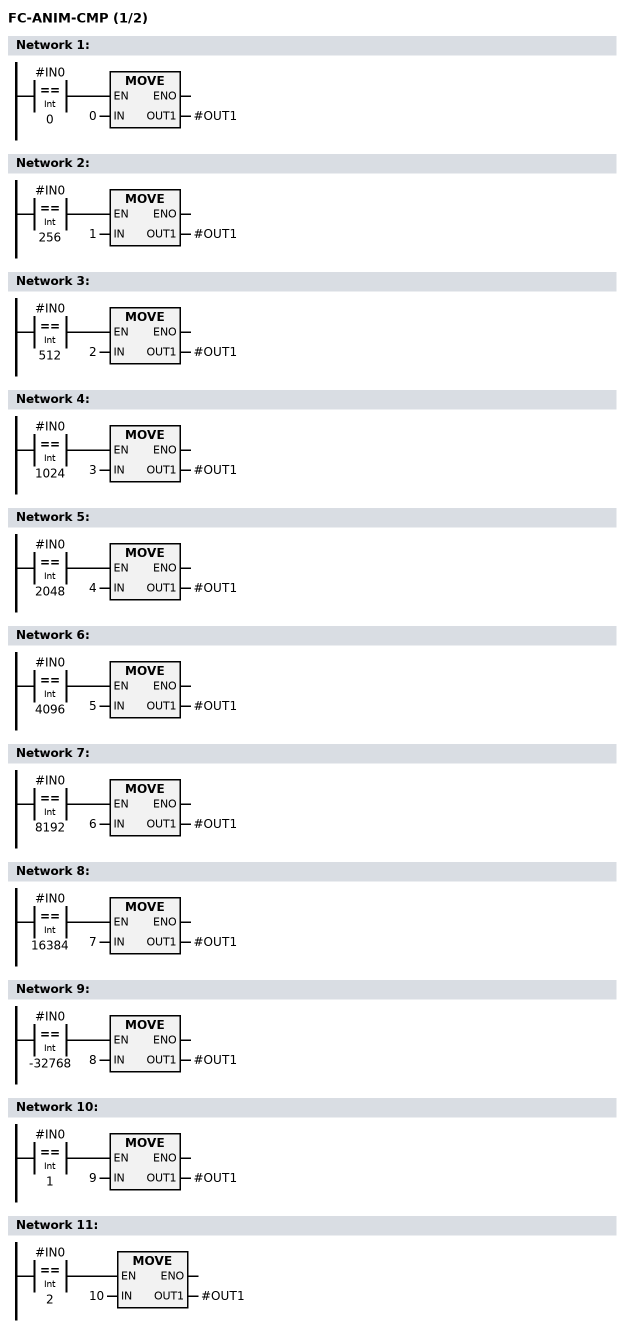
   RUNG wire#powerrail
      { S7_Templates := "SrcType := Int" } EQ_Contact(in1 := #IN0, in2 := 0)
      { S7_GenerateENO := "TRUE" } Move(in := 0, out1 => #OUT1)
   END_RUNG
   // the same network as SCL:
   IF #IN0 = 0 THEN #OUT1 := 0; END_IF;
END_REGION

REGION Network 2
   RUNG wire#powerrail
      { S7_Templates := "SrcType := Int" } EQ_Contact(in1 := #IN0, in2 := 256)
      { S7_GenerateENO := "TRUE" } Move(in := 1, out1 => #OUT1)
   END_RUNG
   // the same network as SCL:
   IF #IN0 = 256 THEN #OUT1 := 1; END_IF;
END_REGION

REGION Network 3
   RUNG wire#powerrail
      { S7_Templates := "SrcType := Int" } EQ_Contact(in1 := #IN0, in2 := 512)
      { S7_GenerateENO := "TRUE" } Move(in := 2, out1 => #OUT1)
   END_RUNG
   // the same network as SCL:
   IF #IN0 = 512 THEN #OUT1 := 2; END_IF;
END_REGION

REGION Network 4
   RUNG wire#powerrail
      { S7_Templates := "SrcType := Int" } EQ_Contact(in1 := #IN0, in2 := 1024)
      { S7_GenerateENO := "TRUE" } Move(in := 3, out1 => #OUT1)
   END_RUNG
   // the same network as SCL:
   IF #IN0 = 1024 THEN #OUT1 := 3; END_IF;
END_REGION

REGION Network 5
   RUNG wire#powerrail
      { S7_Templates := "SrcType := Int" } EQ_Contact(in1 := #IN0, in2 := 2048)
      { S7_GenerateENO := "TRUE" } Move(in := 4, out1 => #OUT1)
   END_RUNG
   // the same network as SCL:
   IF #IN0 = 2048 THEN #OUT1 := 4; END_IF;
END_REGION

REGION Network 6
   RUNG wire#powerrail
      { S7_Templates := "SrcType := Int" } EQ_Contact(in1 := #IN0, in2 := 4096)
      { S7_GenerateENO := "TRUE" } Move(in := 5, out1 => #OUT1)
   END_RUNG
   // the same network as SCL:
   IF #IN0 = 4096 THEN #OUT1 := 5; END_IF;
END_REGION

REGION Network 7
   RUNG wire#powerrail
      { S7_Templates := "SrcType := Int" } EQ_Contact(in1 := #IN0, in2 := 8192)
      { S7_GenerateENO := "TRUE" } Move(in := 6, out1 => #OUT1)
   END_RUNG
   // the same network as SCL:
   IF #IN0 = 8192 THEN #OUT1 := 6; END_IF;
END_REGION

REGION Network 8
   RUNG wire#powerrail
      { S7_Templates := "SrcType := Int" } EQ_Contact(in1 := #IN0, in2 := 16384)
      { S7_GenerateENO := "TRUE" } Move(in := 7, out1 => #OUT1)
   END_RUNG
   // the same network as SCL:
   IF #IN0 = 16384 THEN #OUT1 := 7; END_IF;
END_REGION

REGION Network 9
   RUNG wire#powerrail
      { S7_Templates := "SrcType := Int" } EQ_Contact(in1 := #IN0, in2 := -32768)
      { S7_GenerateENO := "TRUE" } Move(in := 8, out1 => #OUT1)
   END_RUNG
   // the same network as SCL:
   IF #IN0 = (-32768) THEN #OUT1 := 8; END_IF;
END_REGION

REGION Network 10
   RUNG wire#powerrail
      { S7_Templates := "SrcType := Int" } EQ_Contact(in1 := #IN0, in2 := 1)
      { S7_GenerateENO := "TRUE" } Move(in := 9, out1 => #OUT1)
   END_RUNG
   // the same network as SCL:
   IF #IN0 = 1 THEN #OUT1 := 9; END_IF;
END_REGION

REGION Network 11
   RUNG wire#powerrail
      { S7_Templates := "SrcType := Int" } EQ_Contact(in1 := #IN0, in2 := 2)
      { S7_GenerateENO := "TRUE" } Move(in := 10, out1 => #OUT1)
   END_RUNG
   // the same network as SCL:
   IF #IN0 = 2 THEN #OUT1 := 10; END_IF;
END_REGION

REGION Network 12
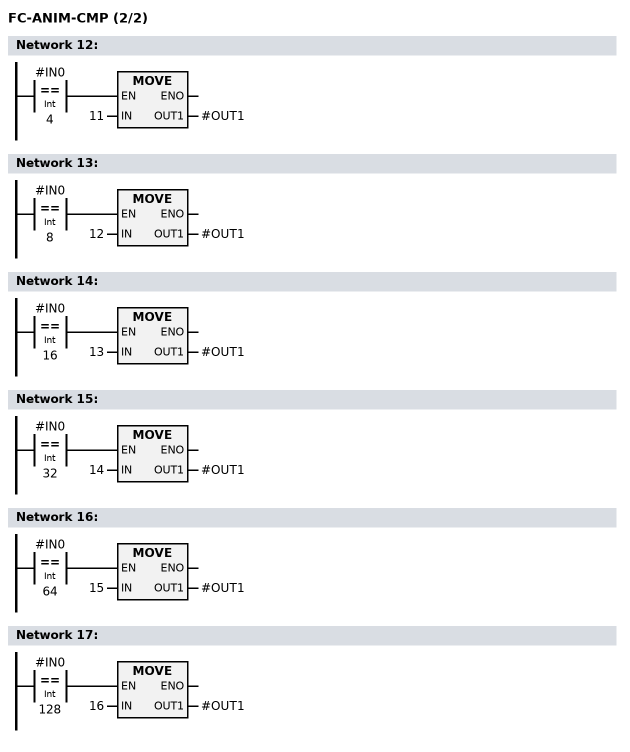
   RUNG wire#powerrail
      { S7_Templates := "SrcType := Int" } EQ_Contact(in1 := #IN0, in2 := 4)
      { S7_GenerateENO := "TRUE" } Move(in := 11, out1 => #OUT1)
   END_RUNG
   // the same network as SCL:
   IF #IN0 = 4 THEN #OUT1 := 11; END_IF;
END_REGION

REGION Network 13
   RUNG wire#powerrail
      { S7_Templates := "SrcType := Int" } EQ_Contact(in1 := #IN0, in2 := 8)
      { S7_GenerateENO := "TRUE" } Move(in := 12, out1 => #OUT1)
   END_RUNG
   // the same network as SCL:
   IF #IN0 = 8 THEN #OUT1 := 12; END_IF;
END_REGION

REGION Network 14
   RUNG wire#powerrail
      { S7_Templates := "SrcType := Int" } EQ_Contact(in1 := #IN0, in2 := 16)
      { S7_GenerateENO := "TRUE" } Move(in := 13, out1 => #OUT1)
   END_RUNG
   // the same network as SCL:
   IF #IN0 = 16 THEN #OUT1 := 13; END_IF;
END_REGION

REGION Network 15
   RUNG wire#powerrail
      { S7_Templates := "SrcType := Int" } EQ_Contact(in1 := #IN0, in2 := 32)
      { S7_GenerateENO := "TRUE" } Move(in := 14, out1 => #OUT1)
   END_RUNG
   // the same network as SCL:
   IF #IN0 = 32 THEN #OUT1 := 14; END_IF;
END_REGION

REGION Network 16
   RUNG wire#powerrail
      { S7_Templates := "SrcType := Int" } EQ_Contact(in1 := #IN0, in2 := 64)
      { S7_GenerateENO := "TRUE" } Move(in := 15, out1 => #OUT1)
   END_RUNG
   // the same network as SCL:
   IF #IN0 = 64 THEN #OUT1 := 15; END_IF;
END_REGION

REGION Network 17
   RUNG wire#powerrail
      { S7_Templates := "SrcType := Int" } EQ_Contact(in1 := #IN0, in2 := 128)
      { S7_GenerateENO := "TRUE" } Move(in := 16, out1 => #OUT1)
   END_RUNG
   // the same network as SCL:
   IF #IN0 = 128 THEN #OUT1 := 16; END_IF;
END_REGION
END_FUNCTION

// folder: Panel/Iluminación

FUNCTION "IluminaciónMTA" : Void   // FC23, LAD
{ S7_Optimized_Access := 'FALSE' }
VERSION : 0.1
// LUC - 05/08/2020
   VAR_TEMP   // added for the SCL form of the ladder/FBD networks
      _s5time1 : S5Time;
   END_VAR
BEGIN

REGION Network 1: Seteo de temporizador desde panel
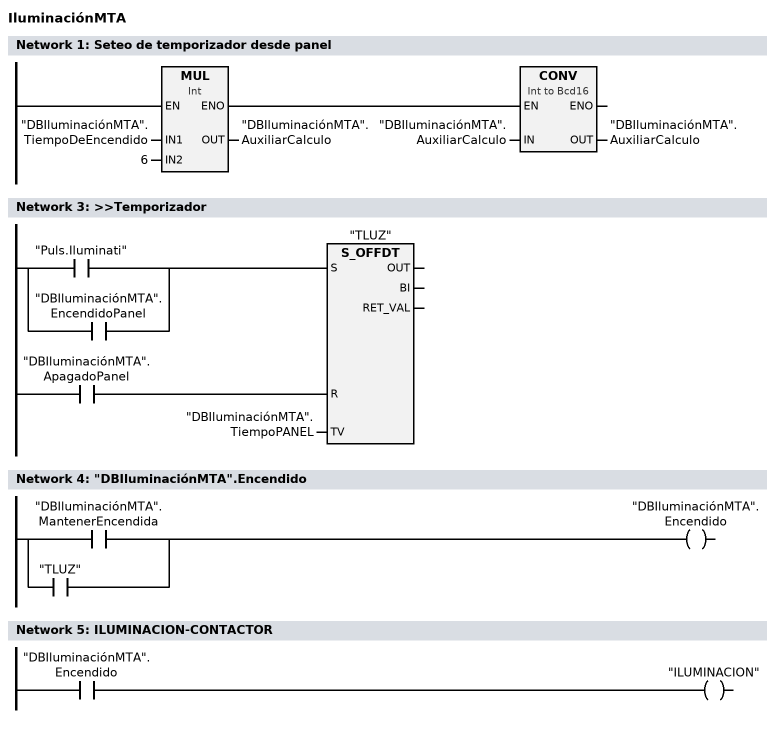
   RUNG wire#powerrail
      { S7_Templates := "SrcType := Int"; S7_GenerateENO := "TRUE" } Mul(in1 := "DBIluminaciónMTA".TiempoDeEncendido, in2 := 6, out => "DBIluminaciónMTA".AuxiliarCalculo)
      { S7_Templates := "[SrcType := Int, DestType := Bcd16]"; S7_GenerateENO := "TRUE" } Convert(in := "DBIluminaciónMTA".AuxiliarCalculo, out => "DBIluminaciónMTA".AuxiliarCalculo)
   END_RUNG
   // the same network as SCL:
   // ENO of a box is taken as its EN; it also drops when the box reports an error
   "DBIluminaciónMTA".AuxiliarCalculo := "DBIluminaciónMTA".TiempoDeEncendido * 6;
   "DBIluminaciónMTA".AuxiliarCalculo := INT_TO_BCD16("DBIluminaciónMTA".AuxiliarCalculo);
END_REGION

REGION Network 2 (STL): Seteo de temporizador desde panel
         L     12288;
         L     "DBIluminaciónMTA".AuxiliarCalculo;
         OW;
         T     "DBIluminaciónMTA".TiempoPANEL;
         NOP   0;
END_REGION

REGION Network 3: >>Temporizador
   RUNG wire#powerrail
      Contact( "Puls.Iluminati" )
      wire#w1
      S_OFFDT(T_NO := "TLUZ", R := wire#w2, TV := "DBIluminaciónMTA".TiempoPANEL, BI =>, RET_VAL =>)
   END_RUNG
   RUNG wire#powerrail
      Contact( "DBIluminaciónMTA".EncendidoPanel )
   END_RUNG wire#w1
   RUNG wire#powerrail
      Contact( "DBIluminaciónMTA".ApagadoPanel )
   END_RUNG wire#w2
   // the same network as SCL:
   #_s5time1 := S_OFFDT(T_NO := "TLUZ",
                        S := "Puls.Iluminati" OR "DBIluminaciónMTA".EncendidoPanel,
                        R := "DBIluminaciónMTA".ApagadoPanel,
                        TV := "DBIluminaciónMTA".TiempoPANEL);
END_REGION

REGION Network 4: "DBIluminaciónMTA".Encendido
   RUNG wire#powerrail
      Contact( "DBIluminaciónMTA".MantenerEncendida )
      wire#w1
      Coil( "DBIluminaciónMTA".Encendido )
   END_RUNG
   RUNG wire#powerrail
      Contact( "TLUZ" )
   END_RUNG wire#w1
   // the same network as SCL:
   "DBIluminaciónMTA".Encendido := "DBIluminaciónMTA".MantenerEncendida OR "TLUZ";
END_REGION

REGION Network 5: ILUMINACION-CONTACTOR
   RUNG wire#powerrail
      Contact( "DBIluminaciónMTA".Encendido )
      Coil( "ILUMINACION" )
   END_RUNG
   // the same network as SCL:
   "ILUMINACION" := "DBIluminaciónMTA".Encendido;
END_REGION
END_FUNCTION

// folder: Secadores/Alta

FUNCTION "EnclavSecAltaMTA" : Void   // FC12, LAD
{ S7_Optimized_Access := 'FALSE' }
VERSION : 0.1
BEGIN

REGION Network 1: Arranque automático MS050
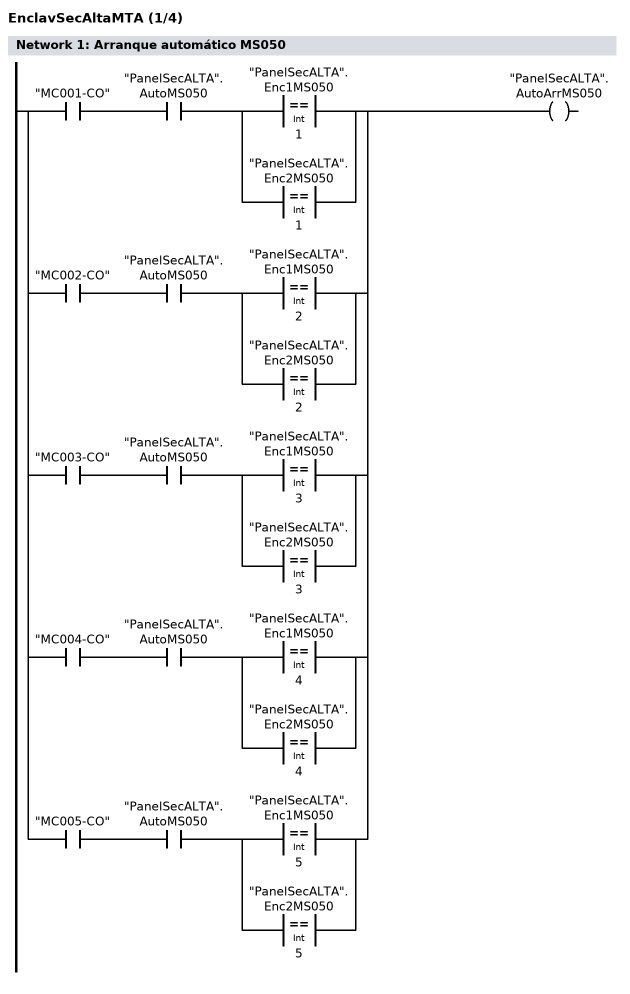
   RUNG wire#powerrail
      Contact( "MC001-CO" )
      Contact( "PanelSecALTA".AutoMS050 )
      wire#w1
      { S7_Templates := "SrcType := Int" } EQ_Contact(in1 := "PanelSecALTA".Enc1MS050, in2 := 1)
      wire#w2
      Coil( "PanelSecALTA".AutoArrMS050 )
   END_RUNG
   RUNG wire#w1
      { S7_Templates := "SrcType := Int" } EQ_Contact(in1 := "PanelSecALTA".Enc2MS050, in2 := 1)
   END_RUNG wire#w2
   RUNG wire#powerrail
      Contact( "MC002-CO" )
      Contact( "PanelSecALTA".AutoMS050 )
      wire#w3
      { S7_Templates := "SrcType := Int" } EQ_Contact(in1 := "PanelSecALTA".Enc1MS050, in2 := 2)
   END_RUNG wire#w2
   RUNG wire#w3
      { S7_Templates := "SrcType := Int" } EQ_Contact(in1 := "PanelSecALTA".Enc2MS050, in2 := 2)
   END_RUNG wire#w2
   RUNG wire#powerrail
      Contact( "MC003-CO" )
      Contact( "PanelSecALTA".AutoMS050 )
      wire#w4
      { S7_Templates := "SrcType := Int" } EQ_Contact(in1 := "PanelSecALTA".Enc1MS050, in2 := 3)
   END_RUNG wire#w2
   RUNG wire#w4
      { S7_Templates := "SrcType := Int" } EQ_Contact(in1 := "PanelSecALTA".Enc2MS050, in2 := 3)
   END_RUNG wire#w2
   RUNG wire#powerrail
      Contact( "MC004-CO" )
      Contact( "PanelSecALTA".AutoMS050 )
      wire#w5
      { S7_Templates := "SrcType := Int" } EQ_Contact(in1 := "PanelSecALTA".Enc1MS050, in2 := 4)
   END_RUNG wire#w2
   RUNG wire#w5
      { S7_Templates := "SrcType := Int" } EQ_Contact(in1 := "PanelSecALTA".Enc2MS050, in2 := 4)
   END_RUNG wire#w2
   RUNG wire#powerrail
      Contact( "MC005-CO" )
      Contact( "PanelSecALTA".AutoMS050 )
      wire#w6
      { S7_Templates := "SrcType := Int" } EQ_Contact(in1 := "PanelSecALTA".Enc1MS050, in2 := 5)
   END_RUNG wire#w2
   RUNG wire#w6
      { S7_Templates := "SrcType := Int" } EQ_Contact(in1 := "PanelSecALTA".Enc2MS050, in2 := 5)
   END_RUNG wire#w2
   // the same network as SCL:
   "PanelSecALTA".AutoArrMS050 := ("MC001-CO" AND "PanelSecALTA".AutoMS050 AND (("PanelSecALTA".Enc1MS050 = 1) OR ("PanelSecALTA".Enc2MS050 = 1))) OR ("MC002-CO" AND "PanelSecALTA".AutoMS050 AND (("PanelSecALTA".Enc1MS050 = 2) OR ("PanelSecALTA".Enc2MS050 = 2))) OR ("MC003-CO" AND "PanelSecALTA".AutoMS050 AND (("PanelSecALTA".Enc1MS050 = 3) OR ("PanelSecALTA".Enc2MS050 = 3))) OR ("MC004-CO" AND "PanelSecALTA".AutoMS050 AND (("PanelSecALTA".Enc1MS050 = 4) OR ("PanelSecALTA".Enc2MS050 = 4))) OR ("MC005-CO" AND "PanelSecALTA".AutoMS050 AND (("PanelSecALTA".Enc1MS050 = 5) OR ("PanelSecALTA".Enc2MS050 = 5)));
END_REGION

REGION Network 2: Arranque automático MS051
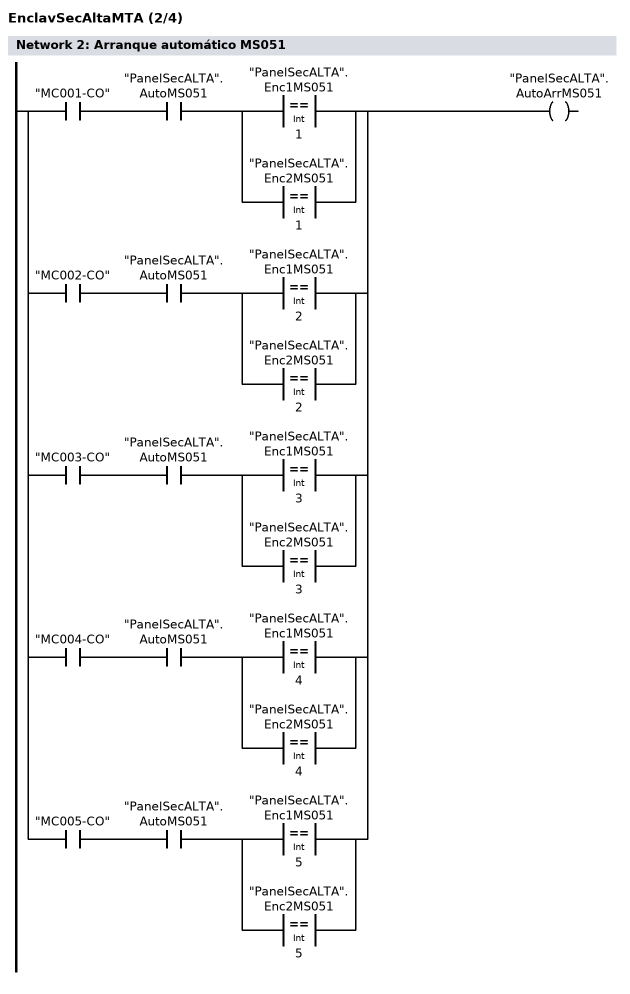
   RUNG wire#powerrail
      Contact( "MC001-CO" )
      Contact( "PanelSecALTA".AutoMS051 )
      wire#w1
      { S7_Templates := "SrcType := Int" } EQ_Contact(in1 := "PanelSecALTA".Enc1MS051, in2 := 1)
      wire#w2
      Coil( "PanelSecALTA".AutoArrMS051 )
   END_RUNG
   RUNG wire#w1
      { S7_Templates := "SrcType := Int" } EQ_Contact(in1 := "PanelSecALTA".Enc2MS051, in2 := 1)
   END_RUNG wire#w2
   RUNG wire#powerrail
      Contact( "MC002-CO" )
      Contact( "PanelSecALTA".AutoMS051 )
      wire#w3
      { S7_Templates := "SrcType := Int" } EQ_Contact(in1 := "PanelSecALTA".Enc1MS051, in2 := 2)
   END_RUNG wire#w2
   RUNG wire#w3
      { S7_Templates := "SrcType := Int" } EQ_Contact(in1 := "PanelSecALTA".Enc2MS051, in2 := 2)
   END_RUNG wire#w2
   RUNG wire#powerrail
      Contact( "MC003-CO" )
      Contact( "PanelSecALTA".AutoMS051 )
      wire#w4
      { S7_Templates := "SrcType := Int" } EQ_Contact(in1 := "PanelSecALTA".Enc1MS051, in2 := 3)
   END_RUNG wire#w2
   RUNG wire#w4
      { S7_Templates := "SrcType := Int" } EQ_Contact(in1 := "PanelSecALTA".Enc2MS051, in2 := 3)
   END_RUNG wire#w2
   RUNG wire#powerrail
      Contact( "MC004-CO" )
      Contact( "PanelSecALTA".AutoMS051 )
      wire#w5
      { S7_Templates := "SrcType := Int" } EQ_Contact(in1 := "PanelSecALTA".Enc1MS051, in2 := 4)
   END_RUNG wire#w2
   RUNG wire#w5
      { S7_Templates := "SrcType := Int" } EQ_Contact(in1 := "PanelSecALTA".Enc2MS051, in2 := 4)
   END_RUNG wire#w2
   RUNG wire#powerrail
      Contact( "MC005-CO" )
      Contact( "PanelSecALTA".AutoMS051 )
      wire#w6
      { S7_Templates := "SrcType := Int" } EQ_Contact(in1 := "PanelSecALTA".Enc1MS051, in2 := 5)
   END_RUNG wire#w2
   RUNG wire#w6
      { S7_Templates := "SrcType := Int" } EQ_Contact(in1 := "PanelSecALTA".Enc2MS051, in2 := 5)
   END_RUNG wire#w2
   // the same network as SCL:
   "PanelSecALTA".AutoArrMS051 := ("MC001-CO" AND "PanelSecALTA".AutoMS051 AND (("PanelSecALTA".Enc1MS051 = 1) OR ("PanelSecALTA".Enc2MS051 = 1))) OR ("MC002-CO" AND "PanelSecALTA".AutoMS051 AND (("PanelSecALTA".Enc1MS051 = 2) OR ("PanelSecALTA".Enc2MS051 = 2))) OR ("MC003-CO" AND "PanelSecALTA".AutoMS051 AND (("PanelSecALTA".Enc1MS051 = 3) OR ("PanelSecALTA".Enc2MS051 = 3))) OR ("MC004-CO" AND "PanelSecALTA".AutoMS051 AND (("PanelSecALTA".Enc1MS051 = 4) OR ("PanelSecALTA".Enc2MS051 = 4))) OR ("MC005-CO" AND "PanelSecALTA".AutoMS051 AND (("PanelSecALTA".Enc1MS051 = 5) OR ("PanelSecALTA".Enc2MS051 = 5)));
END_REGION

REGION Network 3: Arranque automático MS052
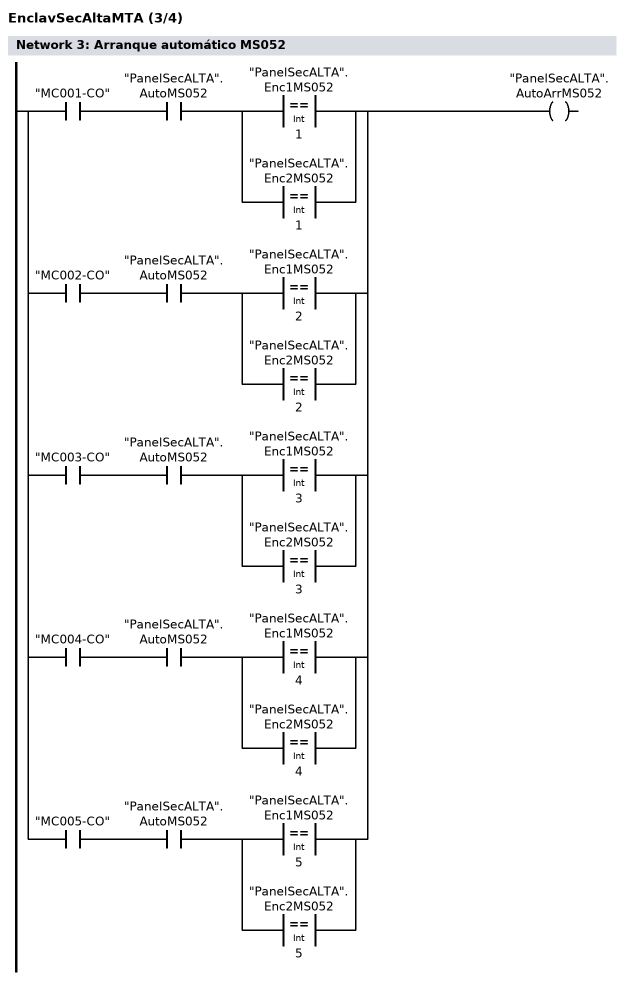
   RUNG wire#powerrail
      Contact( "MC001-CO" )
      Contact( "PanelSecALTA".AutoMS052 )
      wire#w1
      { S7_Templates := "SrcType := Int" } EQ_Contact(in1 := "PanelSecALTA".Enc1MS052, in2 := 1)
      wire#w2
      Coil( "PanelSecALTA".AutoArrMS052 )
   END_RUNG
   RUNG wire#w1
      { S7_Templates := "SrcType := Int" } EQ_Contact(in1 := "PanelSecALTA".Enc2MS052, in2 := 1)
   END_RUNG wire#w2
   RUNG wire#powerrail
      Contact( "MC002-CO" )
      Contact( "PanelSecALTA".AutoMS052 )
      wire#w3
      { S7_Templates := "SrcType := Int" } EQ_Contact(in1 := "PanelSecALTA".Enc1MS052, in2 := 2)
   END_RUNG wire#w2
   RUNG wire#w3
      { S7_Templates := "SrcType := Int" } EQ_Contact(in1 := "PanelSecALTA".Enc2MS052, in2 := 2)
   END_RUNG wire#w2
   RUNG wire#powerrail
      Contact( "MC003-CO" )
      Contact( "PanelSecALTA".AutoMS052 )
      wire#w4
      { S7_Templates := "SrcType := Int" } EQ_Contact(in1 := "PanelSecALTA".Enc1MS052, in2 := 3)
   END_RUNG wire#w2
   RUNG wire#w4
      { S7_Templates := "SrcType := Int" } EQ_Contact(in1 := "PanelSecALTA".Enc2MS052, in2 := 3)
   END_RUNG wire#w2
   RUNG wire#powerrail
      Contact( "MC004-CO" )
      Contact( "PanelSecALTA".AutoMS052 )
      wire#w5
      { S7_Templates := "SrcType := Int" } EQ_Contact(in1 := "PanelSecALTA".Enc1MS052, in2 := 4)
   END_RUNG wire#w2
   RUNG wire#w5
      { S7_Templates := "SrcType := Int" } EQ_Contact(in1 := "PanelSecALTA".Enc2MS052, in2 := 4)
   END_RUNG wire#w2
   RUNG wire#powerrail
      Contact( "MC005-CO" )
      Contact( "PanelSecALTA".AutoMS052 )
      wire#w6
      { S7_Templates := "SrcType := Int" } EQ_Contact(in1 := "PanelSecALTA".Enc1MS052, in2 := 5)
   END_RUNG wire#w2
   RUNG wire#w6
      { S7_Templates := "SrcType := Int" } EQ_Contact(in1 := "PanelSecALTA".Enc2MS052, in2 := 5)
   END_RUNG wire#w2
   // the same network as SCL:
   "PanelSecALTA".AutoArrMS052 := ("MC001-CO" AND "PanelSecALTA".AutoMS052 AND (("PanelSecALTA".Enc1MS052 = 1) OR ("PanelSecALTA".Enc2MS052 = 1))) OR ("MC002-CO" AND "PanelSecALTA".AutoMS052 AND (("PanelSecALTA".Enc1MS052 = 2) OR ("PanelSecALTA".Enc2MS052 = 2))) OR ("MC003-CO" AND "PanelSecALTA".AutoMS052 AND (("PanelSecALTA".Enc1MS052 = 3) OR ("PanelSecALTA".Enc2MS052 = 3))) OR ("MC004-CO" AND "PanelSecALTA".AutoMS052 AND (("PanelSecALTA".Enc1MS052 = 4) OR ("PanelSecALTA".Enc2MS052 = 4))) OR ("MC005-CO" AND "PanelSecALTA".AutoMS052 AND (("PanelSecALTA".Enc1MS052 = 5) OR ("PanelSecALTA".Enc2MS052 = 5)));
END_REGION

REGION Network 4: Arranque automático MS053
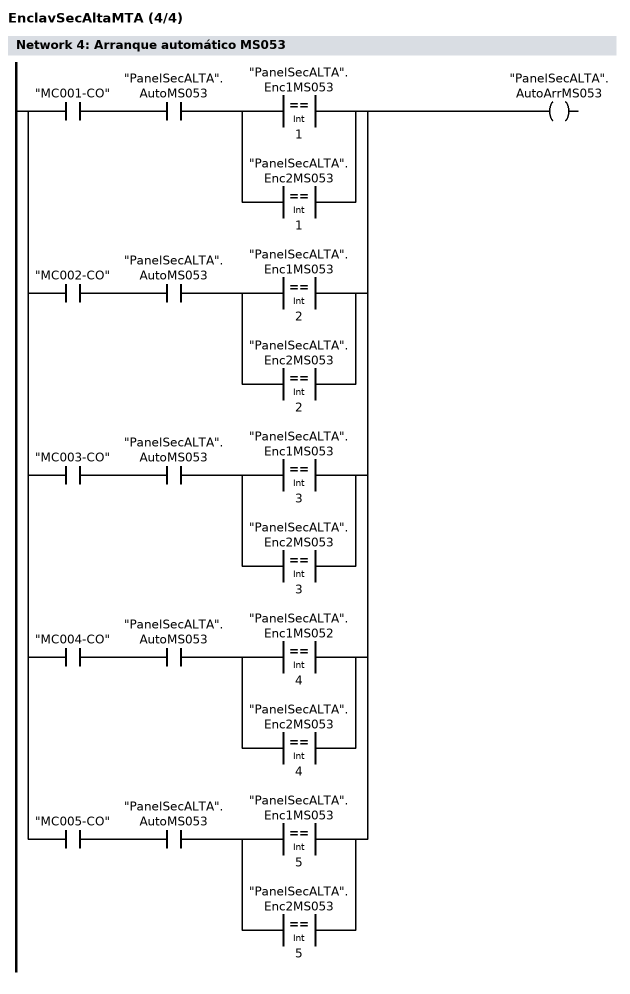
   RUNG wire#powerrail
      Contact( "MC001-CO" )
      Contact( "PanelSecALTA".AutoMS053 )
      wire#w1
      { S7_Templates := "SrcType := Int" } EQ_Contact(in1 := "PanelSecALTA".Enc1MS053, in2 := 1)
      wire#w2
      Coil( "PanelSecALTA".AutoArrMS053 )
   END_RUNG
   RUNG wire#w1
      { S7_Templates := "SrcType := Int" } EQ_Contact(in1 := "PanelSecALTA".Enc2MS053, in2 := 1)
   END_RUNG wire#w2
   RUNG wire#powerrail
      Contact( "MC002-CO" )
      Contact( "PanelSecALTA".AutoMS053 )
      wire#w3
      { S7_Templates := "SrcType := Int" } EQ_Contact(in1 := "PanelSecALTA".Enc1MS053, in2 := 2)
   END_RUNG wire#w2
   RUNG wire#w3
      { S7_Templates := "SrcType := Int" } EQ_Contact(in1 := "PanelSecALTA".Enc2MS053, in2 := 2)
   END_RUNG wire#w2
   RUNG wire#powerrail
      Contact( "MC003-CO" )
      Contact( "PanelSecALTA".AutoMS053 )
      wire#w4
      { S7_Templates := "SrcType := Int" } EQ_Contact(in1 := "PanelSecALTA".Enc1MS053, in2 := 3)
   END_RUNG wire#w2
   RUNG wire#w4
      { S7_Templates := "SrcType := Int" } EQ_Contact(in1 := "PanelSecALTA".Enc2MS053, in2 := 3)
   END_RUNG wire#w2
   RUNG wire#powerrail
      Contact( "MC004-CO" )
      Contact( "PanelSecALTA".AutoMS053 )
      wire#w5
      { S7_Templates := "SrcType := Int" } EQ_Contact(in1 := "PanelSecALTA".Enc1MS052, in2 := 4)
   END_RUNG wire#w2
   RUNG wire#w5
      { S7_Templates := "SrcType := Int" } EQ_Contact(in1 := "PanelSecALTA".Enc2MS053, in2 := 4)
   END_RUNG wire#w2
   RUNG wire#powerrail
      Contact( "MC005-CO" )
      Contact( "PanelSecALTA".AutoMS053 )
      wire#w6
      { S7_Templates := "SrcType := Int" } EQ_Contact(in1 := "PanelSecALTA".Enc1MS053, in2 := 5)
   END_RUNG wire#w2
   RUNG wire#w6
      { S7_Templates := "SrcType := Int" } EQ_Contact(in1 := "PanelSecALTA".Enc2MS053, in2 := 5)
   END_RUNG wire#w2
   // the same network as SCL:
   "PanelSecALTA".AutoArrMS053 := ("MC001-CO" AND "PanelSecALTA".AutoMS053 AND (("PanelSecALTA".Enc1MS053 = 1) OR ("PanelSecALTA".Enc2MS053 = 1))) OR ("MC002-CO" AND "PanelSecALTA".AutoMS053 AND (("PanelSecALTA".Enc1MS053 = 2) OR ("PanelSecALTA".Enc2MS053 = 2))) OR ("MC003-CO" AND "PanelSecALTA".AutoMS053 AND (("PanelSecALTA".Enc1MS053 = 3) OR ("PanelSecALTA".Enc2MS053 = 3))) OR ("MC004-CO" AND "PanelSecALTA".AutoMS053 AND (("PanelSecALTA".Enc1MS052 = 4) OR ("PanelSecALTA".Enc2MS053 = 4))) OR ("MC005-CO" AND "PanelSecALTA".AutoMS053 AND (("PanelSecALTA".Enc1MS053 = 5) OR ("PanelSecALTA".Enc2MS053 = 5)));
END_REGION
END_FUNCTION

// folder: Torres de Agua/Torres Cavaleto

FUNCTION "TorresCavaletoMTA" : Void   // FC14, LAD
{ S7_Optimized_Access := 'FALSE' }
VERSION : 0.1
BEGIN

REGION Network 1: Comandos MV030 / Comandos desde Panel para MV030 - Ventilador 2 Torres de enfriamiento Cavaleto
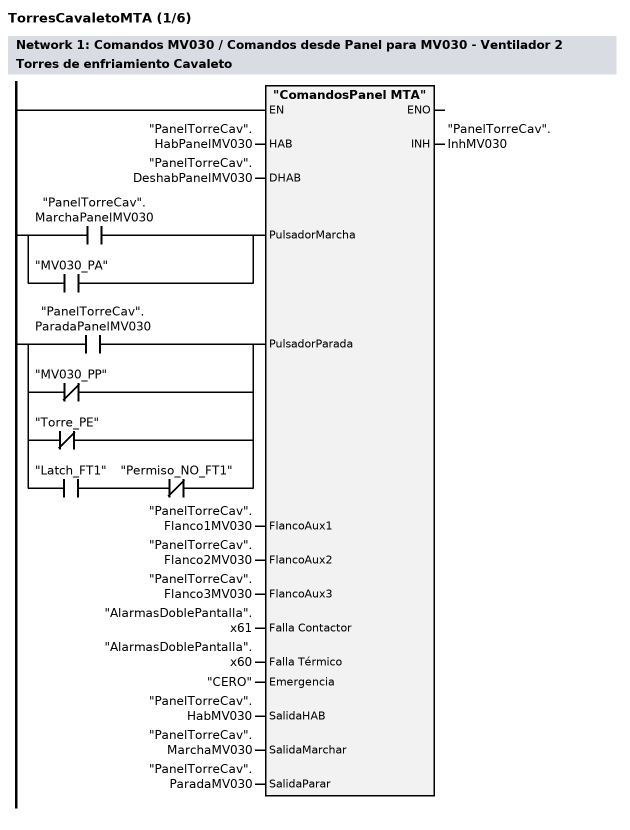
   RUNG wire#powerrail
      "ComandosPanel MTA"(PulsadorMarcha := wire#w1, PulsadorParada := wire#w2, HAB := "PanelTorreCav".HabPanelMV030, DHAB := "PanelTorreCav".DeshabPanelMV030, FlancoAux1 := "PanelTorreCav".Flanco1MV030, FlancoAux2 := "PanelTorreCav".Flanco2MV030, FlancoAux3 := "PanelTorreCav".Flanco3MV030, "Falla Contactor" := "AlarmasDoblePantalla".x61, "Falla Térmico" := "AlarmasDoblePantalla".x60, Emergencia := "CERO", SalidaHAB := "PanelTorreCav".HabMV030, SalidaMarchar := "PanelTorreCav".MarchaMV030, SalidaParar := "PanelTorreCav".ParadaMV030, INH => "PanelTorreCav".InhMV030)
   END_RUNG
   RUNG wire#powerrail
      Contact( "PanelTorreCav".MarchaPanelMV030 )
   END_RUNG wire#w1
   RUNG wire#powerrail
      Contact( "MV030_PA" )
   END_RUNG wire#w1
   RUNG wire#powerrail
      Contact( "PanelTorreCav".ParadaPanelMV030 )
   END_RUNG wire#w2
   RUNG wire#powerrail
      I_Contact( "MV030_PP" )
   END_RUNG wire#w2
   RUNG wire#powerrail
      I_Contact( "Torre_PE" )
   END_RUNG wire#w2
   RUNG wire#powerrail
      Contact( "Latch_FT1" )
      I_Contact( "Permiso_NO_FT1" )
   END_RUNG wire#w2
   // the same network as SCL:
   "ComandosPanel MTA"(HAB := "PanelTorreCav".HabPanelMV030,
                       DHAB := "PanelTorreCav".DeshabPanelMV030,
                       PulsadorMarcha := "PanelTorreCav".MarchaPanelMV030 OR "MV030_PA",
                       PulsadorParada := "PanelTorreCav".ParadaPanelMV030 OR NOT "MV030_PP" OR NOT "Torre_PE" OR ("Latch_FT1" AND NOT "Permiso_NO_FT1"),
                       FlancoAux1 := "PanelTorreCav".Flanco1MV030,
                       FlancoAux2 := "PanelTorreCav".Flanco2MV030,
                       FlancoAux3 := "PanelTorreCav".Flanco3MV030,
                       "Falla Contactor" := "AlarmasDoblePantalla".x61,
                       "Falla Térmico" := "AlarmasDoblePantalla".x60,
                       Emergencia := "CERO",
                       SalidaHAB := "PanelTorreCav".HabMV030,
                       SalidaMarchar := "PanelTorreCav".MarchaMV030,
                       SalidaParar := "PanelTorreCav".ParadaMV030,
                       INH => "PanelTorreCav".InhMV030);
END_REGION

REGION Network 2: Comandos MV031 / Comandos desde Panel para MV031 - Ventilador 1 Torres de enfriamiento Cavaleto
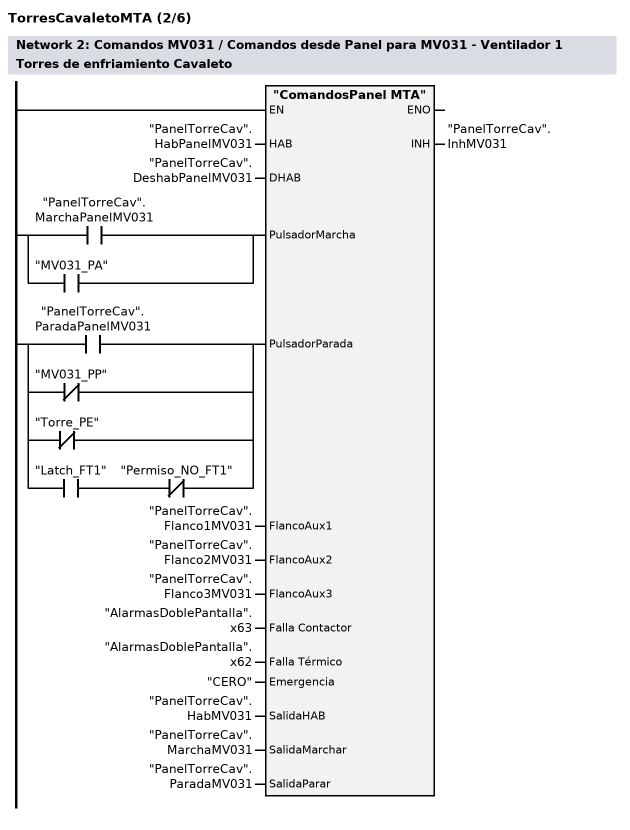
   RUNG wire#powerrail
      "ComandosPanel MTA"(PulsadorMarcha := wire#w1, PulsadorParada := wire#w2, HAB := "PanelTorreCav".HabPanelMV031, DHAB := "PanelTorreCav".DeshabPanelMV031, FlancoAux1 := "PanelTorreCav".Flanco1MV031, FlancoAux2 := "PanelTorreCav".Flanco2MV031, FlancoAux3 := "PanelTorreCav".Flanco3MV031, "Falla Contactor" := "AlarmasDoblePantalla".x63, "Falla Térmico" := "AlarmasDoblePantalla".x62, Emergencia := "CERO", SalidaHAB := "PanelTorreCav".HabMV031, SalidaMarchar := "PanelTorreCav".MarchaMV031, SalidaParar := "PanelTorreCav".ParadaMV031, INH => "PanelTorreCav".InhMV031)
   END_RUNG
   RUNG wire#powerrail
      Contact( "PanelTorreCav".MarchaPanelMV031 )
   END_RUNG wire#w1
   RUNG wire#powerrail
      Contact( "MV031_PA" )
   END_RUNG wire#w1
   RUNG wire#powerrail
      Contact( "PanelTorreCav".ParadaPanelMV031 )
   END_RUNG wire#w2
   RUNG wire#powerrail
      I_Contact( "MV031_PP" )
   END_RUNG wire#w2
   RUNG wire#powerrail
      I_Contact( "Torre_PE" )
   END_RUNG wire#w2
   RUNG wire#powerrail
      Contact( "Latch_FT1" )
      I_Contact( "Permiso_NO_FT1" )
   END_RUNG wire#w2
   // the same network as SCL:
   "ComandosPanel MTA"(HAB := "PanelTorreCav".HabPanelMV031,
                       DHAB := "PanelTorreCav".DeshabPanelMV031,
                       PulsadorMarcha := "PanelTorreCav".MarchaPanelMV031 OR "MV031_PA",
                       PulsadorParada := "PanelTorreCav".ParadaPanelMV031 OR NOT "MV031_PP" OR NOT "Torre_PE" OR ("Latch_FT1" AND NOT "Permiso_NO_FT1"),
                       FlancoAux1 := "PanelTorreCav".Flanco1MV031,
                       FlancoAux2 := "PanelTorreCav".Flanco2MV031,
                       FlancoAux3 := "PanelTorreCav".Flanco3MV031,
                       "Falla Contactor" := "AlarmasDoblePantalla".x63,
                       "Falla Térmico" := "AlarmasDoblePantalla".x62,
                       Emergencia := "CERO",
                       SalidaHAB := "PanelTorreCav".HabMV031,
                       SalidaMarchar := "PanelTorreCav".MarchaMV031,
                       SalidaParar := "PanelTorreCav".ParadaMV031,
                       INH => "PanelTorreCav".InhMV031);
END_REGION

REGION Network 3: Comandos MP014 / Comandos desde Panel para P014 - Bomba 1 Torres de enfriamiento Cavaleto
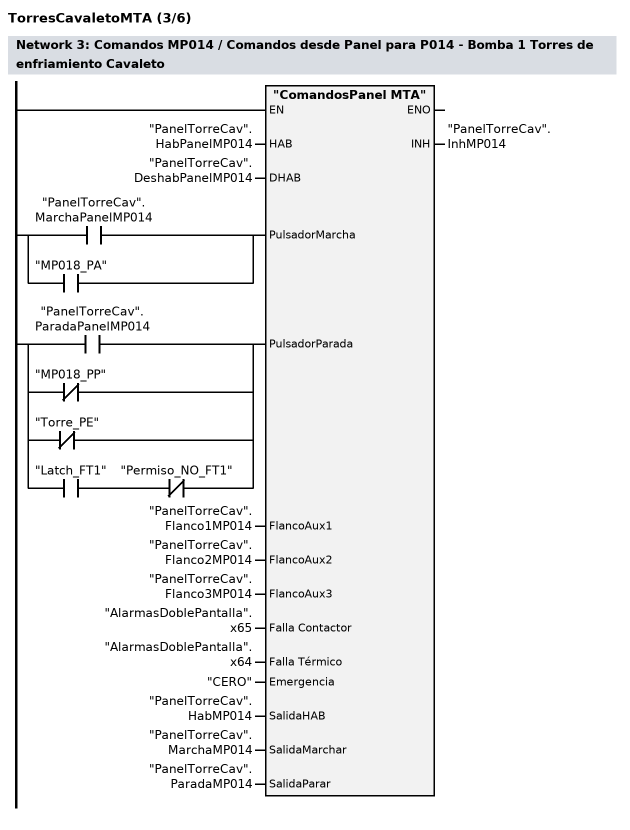
   RUNG wire#powerrail
      "ComandosPanel MTA"(PulsadorMarcha := wire#w1, PulsadorParada := wire#w2, HAB := "PanelTorreCav".HabPanelMP014, DHAB := "PanelTorreCav".DeshabPanelMP014, FlancoAux1 := "PanelTorreCav".Flanco1MP014, FlancoAux2 := "PanelTorreCav".Flanco2MP014, FlancoAux3 := "PanelTorreCav".Flanco3MP014, "Falla Contactor" := "AlarmasDoblePantalla".x65, "Falla Térmico" := "AlarmasDoblePantalla".x64, Emergencia := "CERO", SalidaHAB := "PanelTorreCav".HabMP014, SalidaMarchar := "PanelTorreCav".MarchaMP014, SalidaParar := "PanelTorreCav".ParadaMP014, INH => "PanelTorreCav".InhMP014)
   END_RUNG
   RUNG wire#powerrail
      Contact( "PanelTorreCav".MarchaPanelMP014 )
   END_RUNG wire#w1
   RUNG wire#powerrail
      Contact( "MP018_PA" )
   END_RUNG wire#w1
   RUNG wire#powerrail
      Contact( "PanelTorreCav".ParadaPanelMP014 )
   END_RUNG wire#w2
   RUNG wire#powerrail
      I_Contact( "MP018_PP" )
   END_RUNG wire#w2
   RUNG wire#powerrail
      I_Contact( "Torre_PE" )
   END_RUNG wire#w2
   RUNG wire#powerrail
      Contact( "Latch_FT1" )
      I_Contact( "Permiso_NO_FT1" )
   END_RUNG wire#w2
   // the same network as SCL:
   "ComandosPanel MTA"(HAB := "PanelTorreCav".HabPanelMP014,
                       DHAB := "PanelTorreCav".DeshabPanelMP014,
                       PulsadorMarcha := "PanelTorreCav".MarchaPanelMP014 OR "MP018_PA",
                       PulsadorParada := "PanelTorreCav".ParadaPanelMP014 OR NOT "MP018_PP" OR NOT "Torre_PE" OR ("Latch_FT1" AND NOT "Permiso_NO_FT1"),
                       FlancoAux1 := "PanelTorreCav".Flanco1MP014,
                       FlancoAux2 := "PanelTorreCav".Flanco2MP014,
                       FlancoAux3 := "PanelTorreCav".Flanco3MP014,
                       "Falla Contactor" := "AlarmasDoblePantalla".x65,
                       "Falla Térmico" := "AlarmasDoblePantalla".x64,
                       Emergencia := "CERO",
                       SalidaHAB := "PanelTorreCav".HabMP014,
                       SalidaMarchar := "PanelTorreCav".MarchaMP014,
                       SalidaParar := "PanelTorreCav".ParadaMP014,
                       INH => "PanelTorreCav".InhMP014);
END_REGION

REGION Network 4: Comandos MP015 / Comandos desde Panel para P015 - Bomba 2 Torres de enfriamiento Cavaleto
